// TIA Portal project "uppgift2" (V18)

(* hardware
DEVICE "S7-1500/ET200MP station_1"  S7-1500 station
   slot 0: "Rail_0"  Rack  6ES7 590-1***0-0AA0
   slot 1: "PLC_1"  CPU 1511C-1 PN  6ES7 511-1CK00-0AB0  V2.9
      slot 3: "CPU display_1"  6ES7591-1AA00-0AA0
      slot 32768: "PROFINET interface_1"  X1
         slot 32769: "Port_1"  X1 P1
         slot 32770: "Port_2"  X1 P2
      slot 34817: "Virtual CP interface port_1"  Virtual CP interface port  Virtual CP interface port
DEVICE "HMI_1"  KTP700 Mobile
   slot 0: "HMI_1"  KTP700 Mobile  6AV2 125-2GB03-0AX0  17.0.0.0
   slot 1: "HMI_RT_1"  KTP700 Mobile  6AV2 125-2GB03-0AX0  17.0.0.0
   slot 5: "HMI_1.IE_CP_1"  PROFINET Interface  17.0.0.0
      slot 1: "PROFINET Interface_1"  PROFINET Interface
         slot 1: "Port_1"  Port
*)

// ===== PLC "PLC_1"  CPU 1511C-1 PN =====

VAR_GLOBAL   // PLC tag table "Default tag table"
   "Start Button" AT %I0.0 : Bool;
   "Stop Button" AT %I0.1 : Bool;
   "Reset Button" AT %I0.2 : Bool;
   "Selective Mode" AT %I0.4 : Bool;
   "Base at place" AT %I0.5 : Bool;
   "Lid at place" AT %I0.6 : Bool;
   "Base is clamped" AT %I0.7 : Bool;
   "Lid is clamped" AT %I1.0 : Bool;
   "Item detected" AT %I1.1 : Bool;
   "Part is leaving (Sensor)" AT %I1.2 : Bool;
   "FACTORY I/O (Running)" AT %I1.3 : Bool;
   "Move X (Extend)" AT %Q0.0 : Bool;
   "Move Z (Lower)" AT %Q0.1 : Bool;
   "Grab Item" AT %Q0.2 : Bool;
   "Clamp base" AT %Q0.3 : Bool;
   "Clamp lid" AT %Q0.4 : Bool;
   "Lids emitter" AT %Q0.5 : Bool;
   "Lift Bases Clamp" AT %Q0.6 : Bool;
   "Lift Lids Clamp" AT %Q0.7 : Bool;
   "Counter" AT %QD30 : DInt;
   "Bases Vision Sensor" AT %ID30 : DInt;
   "Lids Vision Sensor" AT %ID34 : DInt;
   "Start Light" AT %Q1.0 : Bool;
   "Stop Light" AT %Q1.1 : Bool;
   "Reset Light" AT %Q1.2 : Bool;
   "Lids conveyor" AT %Q1.3 : Bool;
   "Bases conveyor" AT %Q1.4 : Bool;
   "Bases emitter" AT %Q1.5 : Bool;
   "flanker" AT %I2.4 : Bool;
   "Moving X (Sensor)" AT %I1.4 : Bool;
   "Moving Z (Sensor)" AT %I1.5 : Bool;
   "hmistop" AT %I2.2 : Bool;
   "hmireset" AT %I2.3 : Bool;
   "countyfinalflank" AT %I2.5 : Bool;
   "lids lift clamp limit" AT %I1.6 : Bool;
   "baselift clamp limit" AT %I1.7 : Bool;
   "countyflank" AT %I2.6 : Bool;
END_VAR

// folder: System blocks/Program resources

DATA_BLOCK "IEC_Timer_0_DB"   // DB3
{ S7_Optimized_Access := 'TRUE' }
AUTHOR : Simatic
FAMILY : IEC
NAME : IEC_TMR
VERSION : 1.0
// stored: InstanceOfName IEC_TIMER
"IEC_TIMER"
BEGIN
END_DATA_BLOCK

DATA_BLOCK "IEC_Timer_1_DB"   // DB4
{ S7_Optimized_Access := 'TRUE' }
AUTHOR : Simatic
FAMILY : IEC
NAME : IEC_TMR
VERSION : 1.0
// stored: InstanceOfName IEC_TIMER
"IEC_TIMER"
BEGIN
END_DATA_BLOCK

DATA_BLOCK "IEC_Counter_0_DB_2"   // DB5
{ S7_Optimized_Access := 'TRUE' }
AUTHOR : Simatic
FAMILY : IEC
NAME : CNTR
VERSION : 1.0
// stored: InstanceOfName IEC_COUNTER
"IEC_COUNTER"
BEGIN
END_DATA_BLOCK

DATA_BLOCK "IEC_Timer_0_DB_2"   // DB6
{ S7_Optimized_Access := 'TRUE' }
AUTHOR : Simatic
FAMILY : IEC
NAME : IEC_TMR
VERSION : 1.0
// stored: InstanceOfName IEC_TIMER
"IEC_TIMER"
BEGIN
END_DATA_BLOCK

DATA_BLOCK "IEC_Counter_0_DB_3"   // DB8
{ S7_Optimized_Access := 'TRUE' }
AUTHOR : Simatic
FAMILY : IEC
NAME : CNTR
VERSION : 1.0
// stored: InstanceOfName IEC_COUNTER
"IEC_COUNTER"
BEGIN
END_DATA_BLOCK

DATA_BLOCK "IEC_Counter_0_DB_4"   // DB10
{ S7_Optimized_Access := 'TRUE' }
AUTHOR : Simatic
FAMILY : IEC
NAME : CNTR
VERSION : 1.0
// stored: InstanceOfName IEC_COUNTER
"IEC_COUNTER"
BEGIN
END_DATA_BLOCK

DATA_BLOCK "IEC_Counter_0_DB_6"   // DB11
{ S7_Optimized_Access := 'TRUE' }
AUTHOR : Simatic
FAMILY : IEC
NAME : CNTR
VERSION : 1.0
// stored: InstanceOfName IEC_COUNTER
"IEC_COUNTER"
BEGIN
END_DATA_BLOCK

DATA_BLOCK "IEC_Counter_1_DB_1"   // DB12
{ S7_Optimized_Access := 'TRUE' }
AUTHOR : Simatic
FAMILY : IEC
NAME : CNTR
VERSION : 1.0
// stored: InstanceOfName IEC_COUNTER
"IEC_COUNTER"
BEGIN
END_DATA_BLOCK

DATA_BLOCK "IEC_Counter_0_DB_7"   // DB13
{ S7_Optimized_Access := 'TRUE' }
AUTHOR : Simatic
FAMILY : IEC
NAME : CNTR
VERSION : 1.0
// stored: InstanceOfName IEC_COUNTER
"IEC_COUNTER"
BEGIN
END_DATA_BLOCK

DATA_BLOCK "IEC_Counter_0_DB_5"   // DB14
{ S7_Optimized_Access := 'TRUE' }
AUTHOR : Simatic
FAMILY : IEC
NAME : CNTR
VERSION : 1.0
// stored: InstanceOfName IEC_COUNTER
"IEC_COUNTER"
BEGIN
END_DATA_BLOCK

DATA_BLOCK "IEC_Counter_0_DB_8"   // DB15
{ S7_Optimized_Access := 'TRUE' }
AUTHOR : Simatic
FAMILY : IEC
NAME : CNTR
VERSION : 1.0
// stored: InstanceOfName IEC_COUNTER
"IEC_COUNTER"
BEGIN
END_DATA_BLOCK

DATA_BLOCK "IEC_Counter_0_DB_9"   // DB16
{ S7_Optimized_Access := 'TRUE' }
AUTHOR : Simatic
FAMILY : IEC
NAME : CNTR
VERSION : 1.0
// stored: InstanceOfName IEC_COUNTER
"IEC_COUNTER"
BEGIN
END_DATA_BLOCK

DATA_BLOCK "IEC_Timer_5_DB"   // DB17
{ S7_Optimized_Access := 'TRUE' }
AUTHOR : Simatic
FAMILY : IEC
NAME : IEC_TMR
VERSION : 1.0
// stored: InstanceOfName IEC_TIMER
"IEC_TIMER"
BEGIN
END_DATA_BLOCK

DATA_BLOCK "IEC_Counter_0_DB"   // DB18
{ S7_Optimized_Access := 'TRUE' }
AUTHOR : Simatic
FAMILY : IEC
NAME : CNTR
VERSION : 1.0
// stored: InstanceOfName IEC_COUNTER
"IEC_COUNTER"
BEGIN
END_DATA_BLOCK

DATA_BLOCK "IEC_Timer_0_DB_4"   // DB20
{ S7_Optimized_Access := 'TRUE' }
AUTHOR : Simatic
FAMILY : IEC
NAME : IEC_TMR
VERSION : 1.0
// stored: InstanceOfName IEC_TIMER
"IEC_TIMER"
BEGIN
END_DATA_BLOCK

// folder: databases

DATA_BLOCK "outputs"   // DB1
{ S7_Optimized_Access := 'TRUE' }
VERSION : 0.1
   VAR
      RESETBUTTONHMI : Bool;
      Acutators : Struct
         "Move X (Extend)" : Bool;
         "Move Z (Lower)" : Bool;
         "Grab Item" : Bool;
         "Clamp base" : Bool;
         "Clamp lid" : Bool;
         "Lift Bases Clamp" : Bool;
         "Lift Lids Clamp" : Bool;
      END_STRUCT;
      BoxesCounters : Struct
         "green lids" : Int;
         "green bases" : Int;
         "blue lids" : Int;
         "blue bases" : Int;
         "bluegreen box" : Int;   // blå lock grön bas
         "greenblue box" : Int;   // grön bas blå lock
         "blue boxs" : Int;
         "green boxs" : Int;
         totalpartscounter : Int;
      END_STRUCT;
      Checks : Struct
         isreset : Bool;
         selectivestmode : Bool;
         pauseforselective : Bool;
      END_STRUCT;
      Modes : Struct
         "Run mode" : Bool;
         "Reset mode" : Bool;
         "Stop mode" : Bool;
      END_STRUCT;
      "Hmi-Producer" : Struct
         producedboxes : Int;
         toproduce : Int := 0;
      END_STRUCT;
   END_VAR
BEGIN
END_DATA_BLOCK

DATA_BLOCK "inputs"   // DB2
{ S7_Optimized_Access := 'TRUE' }
VERSION : 0.1
   VAR
      buttons : Struct
         "Start Button" : Bool;
         "Stop Button" : Bool;
         "Reset Button" : Bool;
      END_STRUCT;
      Sensors : Struct
         "Item detected" : Bool;
         "lid sensor value" : DInt;
      END_STRUCT;
      Sequences : Struct
         insequence : DInt;
         basesecquence : DInt;
         robotarmsequence : DInt;
      END_STRUCT;
      "green light" : Bool;
   END_VAR
BEGIN
END_DATA_BLOCK

DATA_BLOCK "functiondatabase"   // DB9
{ S7_Optimized_Access := 'TRUE' }
VERSION : 0.1
// stored: InstanceOfName hmi-order-limit&Color-total
"hmi-order-limit&Color-total"
BEGIN
END_DATA_BLOCK

DATA_BLOCK "tondb"   // DB19
{ S7_Optimized_Access := 'TRUE' }
VERSION : 0.1
   VAR
      IN : Bool;
      PT : Time := T#7000ms;
      Q : Bool;
      ET : Time;
   END_VAR
BEGIN
END_DATA_BLOCK

DATA_BLOCK "HMI-DB"   // DB1000
{ S7_Optimized_Access := 'TRUE' }
VERSION : 0.1
   VAR
      Inputs : Struct
         StartLight : Bool;
         StopLight : Bool;
         ResetLight : Bool;
      END_STRUCT;
      "Jogging&Priority" : Struct
         jogmode : Bool;
         hasbeenjogging : Bool;
         "jog bools" : Struct   // hmi jog bools
            "move x" : Bool;
            "move y" : Bool;
            "grab item" : Bool;
            "clamp lid" : Bool;
            "clamp base" : Bool;
            "lift base" : Bool;
            "lift lid" : Bool;
            "lid conv" : Bool;
            "base conv" : Bool;
            lampor : Bool;
         END_STRUCT;
         hmipriority : Bool;
         hmiprioritystate : Bool;
         resetdelivered : Bool;
      END_STRUCT;
   END_VAR
BEGIN
END_DATA_BLOCK

// folder: (top level)

FUNCTION_BLOCK "hmi-order-limit&Color-total"   // FB1, LAD
{ S7_Optimized_Access := 'TRUE' }
VERSION : 0.1
   VAR_OUTPUT
      basesadder : Int;
      lidadder : Int;
   END_VAR
BEGIN

REGION Network 1
   // limits the hmi to produce max 1000
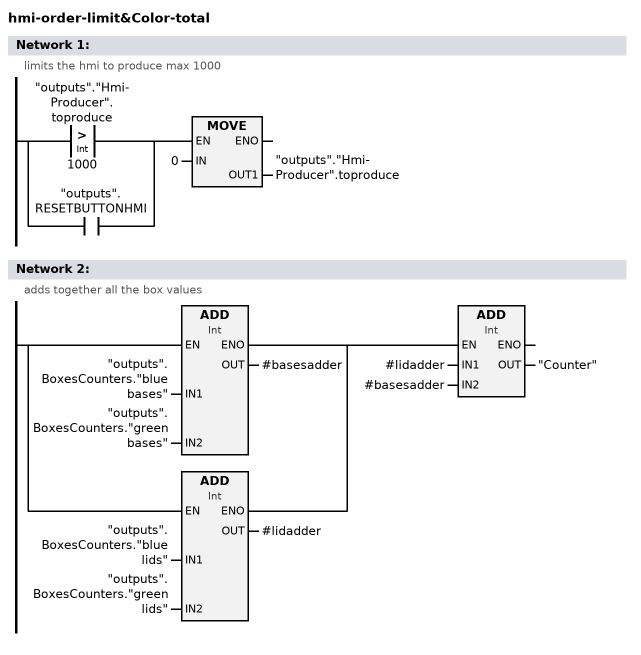
   RUNG wire#powerrail
      { S7_Templates := "SrcType := Int" } GT_Contact(in1 := "outputs"."Hmi-Producer".toproduce, in2 := 1000)
      wire#w1
      Move(in := 0, out1 => "outputs"."Hmi-Producer".toproduce)
   END_RUNG
   RUNG wire#powerrail
      Contact( "outputs".RESETBUTTONHMI )
   END_RUNG wire#w1
   // the same network as SCL:
   IF ("outputs"."Hmi-Producer".toproduce > 1000) OR "outputs".RESETBUTTONHMI THEN
       "outputs"."Hmi-Producer".toproduce := 0;
   END_IF;
END_REGION

REGION Network 2
   // adds together all the box values
   RUNG wire#powerrail
      { S7_Templates := "SrcType := Int" } Add(in1 := "outputs".BoxesCounters."blue bases", in2 := "outputs".BoxesCounters."green bases", out => #basesadder)
      wire#w1
      { S7_Templates := "SrcType := Int" } Add(in1 := #lidadder, in2 := #basesadder, out => "Counter")
   END_RUNG
   RUNG wire#powerrail
      { S7_Templates := "SrcType := Int" } Add(in1 := "outputs".BoxesCounters."blue lids", in2 := "outputs".BoxesCounters."green lids", out => #lidadder)
   END_RUNG wire#w1
   // the same network as SCL:
   #basesadder := "outputs".BoxesCounters."blue bases" + "outputs".BoxesCounters."green bases";
   #lidadder := "outputs".BoxesCounters."blue lids" + "outputs".BoxesCounters."green lids";
   IF TRUE OR TRUE THEN "Counter" := #lidadder + #basesadder; END_IF;
END_REGION
END_FUNCTION_BLOCK

FUNCTION "robotarm" : Void   // FC5, LAD
{ S7_Optimized_Access := 'TRUE' }
VERSION : 0.1
   VAR_TEMP   // added for the SCL form of the ladder/FBD networks
      _w1 : Bool;
   END_VAR
BEGIN

REGION Network 1
   // Both sequence 1 and 3 runs in the same network in an "or" statement, because both sequences need to use the "move z" acutator.
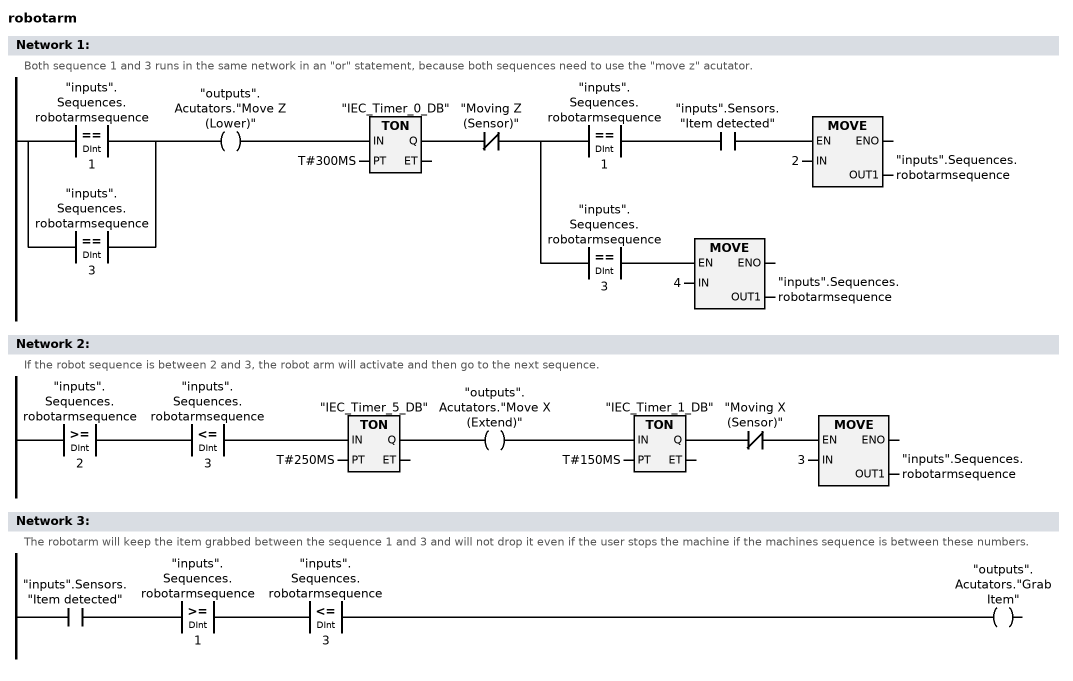
   "outputs".Acutators."Move Z (Lower)" := ("inputs".Sequences.robotarmsequence = 1) OR ("inputs".Sequences.robotarmsequence = 3);
   "IEC_Timer_0_DB".TON(IN := "outputs".Acutators."Move Z (Lower)", PT := T#300MS);
   #_w1 := "IEC_Timer_0_DB".Q AND NOT "Moving Z (Sensor)";
   IF #_w1 AND ("inputs".Sequences.robotarmsequence = 1) AND "inputs".Sensors."Item detected" THEN
       "inputs".Sequences.robotarmsequence := 2;
   END_IF;
   IF #_w1 AND ("inputs".Sequences.robotarmsequence = 3) THEN
       "inputs".Sequences.robotarmsequence := 4;
   END_IF;
END_REGION

REGION Network 2
   // If the robot sequence is between 2 and 3, the robot arm will activate and then go to the next sequence.
   "IEC_Timer_5_DB".TON(IN := ("inputs".Sequences.robotarmsequence >= 2) AND ("inputs".Sequences.robotarmsequence <= 3),
                        PT := T#250MS);
   "outputs".Acutators."Move X (Extend)" := "IEC_Timer_5_DB".Q;
   "IEC_Timer_1_DB".TON(IN := "IEC_Timer_5_DB".Q, PT := T#150MS);
   IF "IEC_Timer_1_DB".Q AND NOT "Moving X (Sensor)" THEN "inputs".Sequences.robotarmsequence := 3; END_IF;
END_REGION

REGION Network 3
   // The robotarm will keep the item grabbed between the sequence 1 and 3 and will not drop it even if the user stops the machine if the machines sequence is between these numbers.
   RUNG wire#powerrail
      Contact( "inputs".Sensors."Item detected" )
      { S7_Templates := "SrcType := DInt" } GE_Contact(in1 := "inputs".Sequences.robotarmsequence, in2 := 1)
      { S7_Templates := "SrcType := DInt" } LE_Contact(in1 := "inputs".Sequences.robotarmsequence, in2 := 3)
      Coil( "outputs".Acutators."Grab Item" )
   END_RUNG
   // the same network as SCL:
   "outputs".Acutators."Grab Item" := "inputs".Sensors."Item detected" AND ("inputs".Sequences.robotarmsequence >= 1) AND ("inputs".Sequences.robotarmsequence <= 3);
END_REGION
END_FUNCTION

FUNCTION "countcolors" : Void   // FC8, LAD
{ S7_Optimized_Access := 'TRUE' }
VERSION : 0.1
// This function counts the colors that passes through the colors sensors, both lid and base and then counts up accordingdly to which color that passed through the sensor.
   VAR_TEMP   // added for the SCL form of the ladder/FBD networks
      _w1 : Bool;
   END_VAR
BEGIN

REGION Network 1: counts final product
   // Counts the total boxes produced.
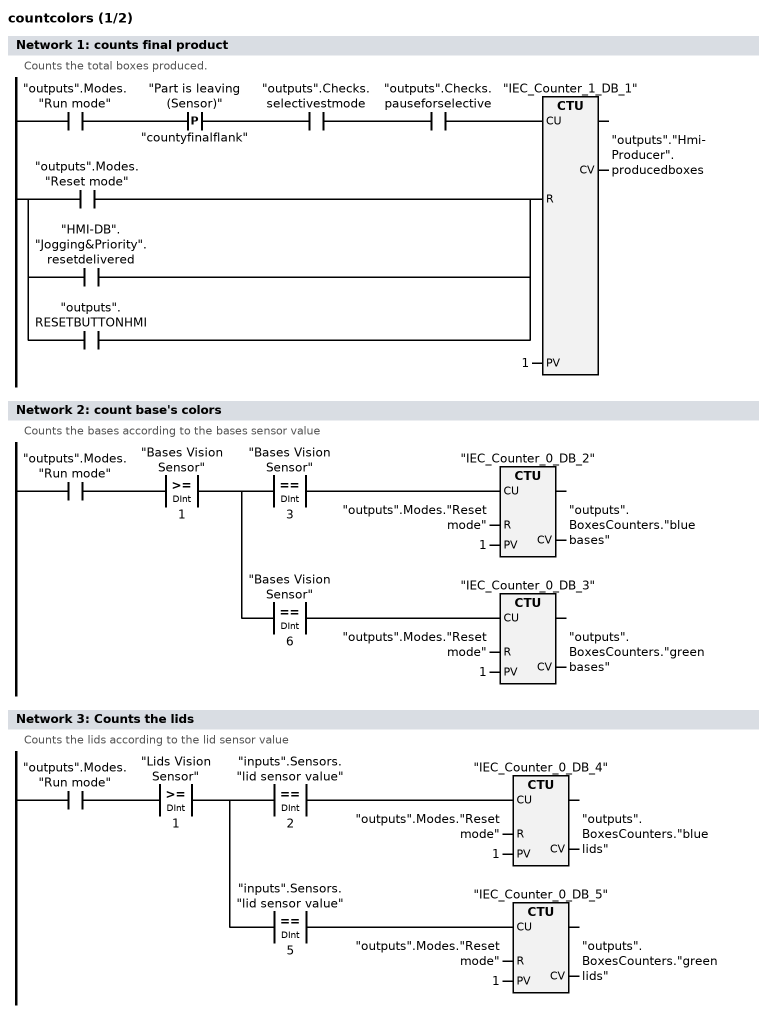
   #_w1 := "outputs".Modes."Run mode" AND "Part is leaving (Sensor)" AND NOT "countyfinalflank";   // rising edge of "Part is leaving (Sensor)"
   "countyfinalflank" := "Part is leaving (Sensor)";
   "IEC_Counter_1_DB_1".CTU(CU := #_w1 AND "outputs".Checks.selectivestmode AND "outputs".Checks.pauseforselective,
                           R := "outputs".Modes."Reset mode" OR "HMI-DB"."Jogging&Priority".resetdelivered OR "outputs".RESETBUTTONHMI,
                           PV := 1,
                           CV => "outputs"."Hmi-Producer".producedboxes);
END_REGION

REGION Network 2: count base's colors
   // Counts the bases according to the bases sensor value
   #_w1 := "outputs".Modes."Run mode" AND ("Bases Vision Sensor" >= 1);
   "IEC_Counter_0_DB_2".CTU(CU := #_w1 AND ("Bases Vision Sensor" = 3),
                           R := "outputs".Modes."Reset mode",
                           PV := 1,
                           CV => "outputs".BoxesCounters."blue bases");
   "IEC_Counter_0_DB_3".CTU(CU := #_w1 AND ("Bases Vision Sensor" = 6),
                           R := "outputs".Modes."Reset mode",
                           PV := 1,
                           CV => "outputs".BoxesCounters."green bases");
END_REGION

REGION Network 3: Counts the lids
   // Counts the lids according to the lid sensor value
   #_w1 := "outputs".Modes."Run mode" AND ("Lids Vision Sensor" >= 1);
   "IEC_Counter_0_DB_4".CTU(CU := #_w1 AND ("inputs".Sensors."lid sensor value" = 2),
                           R := "outputs".Modes."Reset mode",
                           PV := 1,
                           CV => "outputs".BoxesCounters."blue lids");
   "IEC_Counter_0_DB_5".CTU(CU := #_w1 AND ("inputs".Sensors."lid sensor value" = 5),
                           R := "outputs".Modes."Reset mode",
                           PV := 1,
                           CV => "outputs".BoxesCounters."green lids");
END_REGION

REGION Network 4
   // counts if the base and the lid is different colors
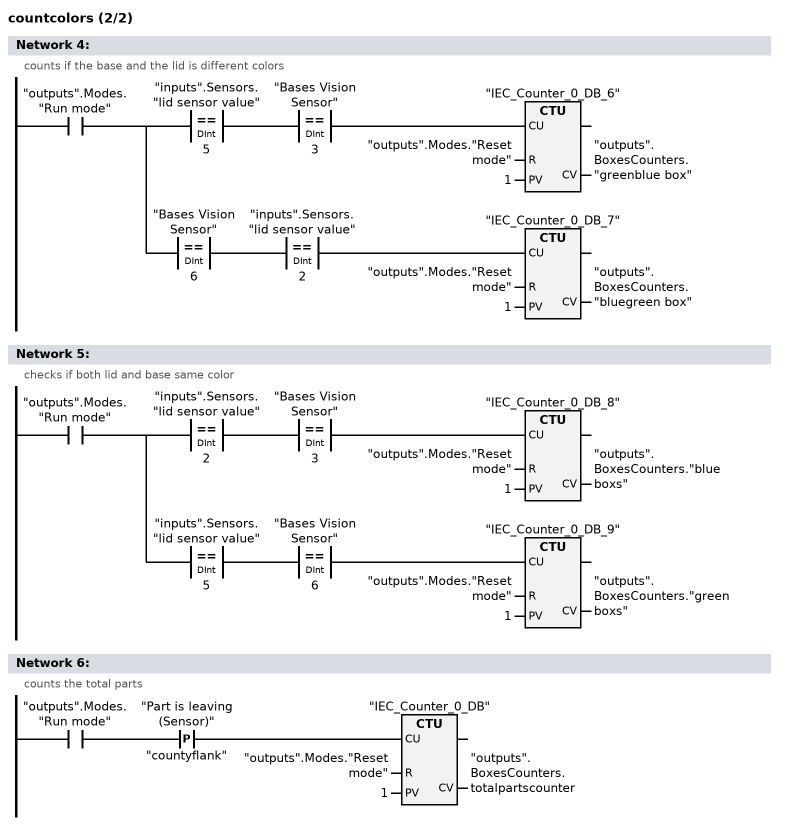
   "IEC_Counter_0_DB_6".CTU(CU := "outputs".Modes."Run mode" AND ("inputs".Sensors."lid sensor value" = 5) AND ("Bases Vision Sensor" = 3),
                           R := "outputs".Modes."Reset mode",
                           PV := 1,
                           CV => "outputs".BoxesCounters."greenblue box");
   "IEC_Counter_0_DB_7".CTU(CU := "outputs".Modes."Run mode" AND ("Bases Vision Sensor" = 6) AND ("inputs".Sensors."lid sensor value" = 2),
                           R := "outputs".Modes."Reset mode",
                           PV := 1,
                           CV => "outputs".BoxesCounters."bluegreen box");
END_REGION

REGION Network 5
   // checks if both lid and base same color
   "IEC_Counter_0_DB_8".CTU(CU := "outputs".Modes."Run mode" AND ("inputs".Sensors."lid sensor value" = 2) AND ("Bases Vision Sensor" = 3),
                           R := "outputs".Modes."Reset mode",
                           PV := 1,
                           CV => "outputs".BoxesCounters."blue boxs");
   "IEC_Counter_0_DB_9".CTU(CU := "outputs".Modes."Run mode" AND ("inputs".Sensors."lid sensor value" = 5) AND ("Bases Vision Sensor" = 6),
                           R := "outputs".Modes."Reset mode",
                           PV := 1,
                           CV => "outputs".BoxesCounters."green boxs");
END_REGION

REGION Network 6
   // counts the total parts
   #_w1 := "outputs".Modes."Run mode" AND "Part is leaving (Sensor)" AND NOT "countyflank";   // rising edge of "Part is leaving (Sensor)"
   "countyflank" := "Part is leaving (Sensor)";
   "IEC_Counter_0_DB".CTU(CU := #_w1,
                          R := "outputs".Modes."Reset mode",
                          PV := 1,
                          CV => "outputs".BoxesCounters.totalpartscounter);
END_REGION
END_FUNCTION

FUNCTION "resetscl" : Void   // FC9, SCL
{ S7_Optimized_Access := 'TRUE' }
VERSION : 0.1
BEGIN


   IF "outputs".Modes."Reset mode" THEN //Checks if its in reset mode
       "inputs".Sequences.basesecquence := 0; //Resets basesequence
       "inputs".Sequences.insequence := 0; //Resets lidsequence

       "tondb".IN := 1; 


       "IEC_Timer_0_DB_4".TON(IN := "tondb".IN, //Timer
                              PT := "tondb".PT,
                              Q => "tondb".Q,
                              ET => "tondb".ET);
       IF "tondb".Q THEN //When timer done then disable reset mode and set "isreset" variable to true
           "outputs".Checks.isreset := 1;
           "outputs".Modes."Reset mode" := 0;

           RESET_TIMER("IEC_Timer_0_DB_4");

       END_IF;

       IF NOT "Item detected" THEN //If arm not holding lid then reset the robot arm sequence
           "inputs".Sequences.robotarmsequence := 0;
       END_IF;

   END_IF;
END_FUNCTION

ORGANIZATION_BLOCK "Main"   // OB1, LAD, ProgramCycle
TITLE = "Main Program Sweep (Cycle)"
{ S7_Optimized_Access := 'TRUE' }
VERSION : 0.1
   VAR_INPUT
      Initial_Call : Bool;   // Initial call of this OB
      Remanence : Bool;   // =True, if remanent data are available
   END_VAR
BEGIN

REGION Network 1
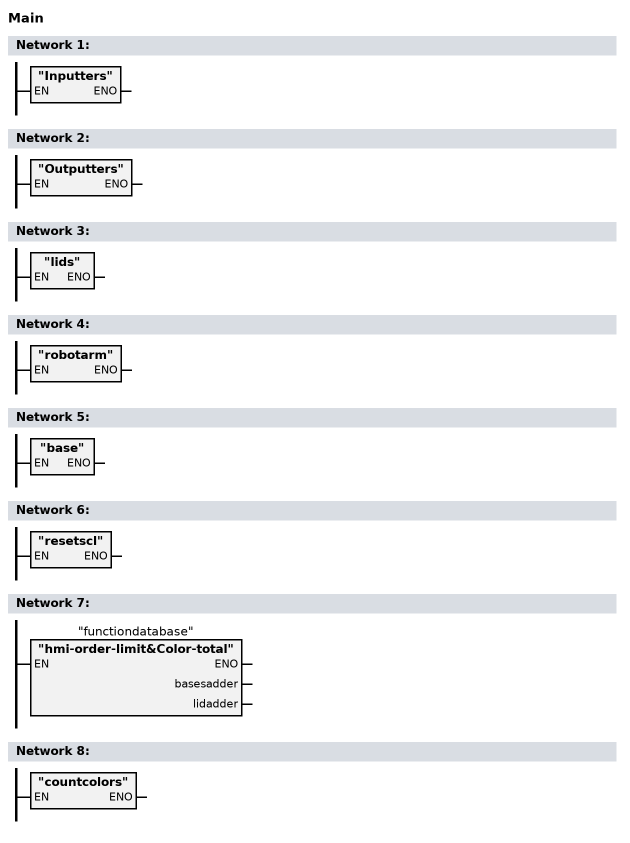
   RUNG wire#powerrail
      "Inputters"()
   END_RUNG
   // the same network as SCL:
   "Inputters"();
END_REGION

REGION Network 2
   RUNG wire#powerrail
      "Outputters"()
   END_RUNG
   // the same network as SCL:
   "Outputters"();
END_REGION

REGION Network 3
   RUNG wire#powerrail
      "lids"()
   END_RUNG
   // the same network as SCL:
   "lids"();
END_REGION

REGION Network 4
   RUNG wire#powerrail
      "robotarm"()
   END_RUNG
   // the same network as SCL:
   "robotarm"();
END_REGION

REGION Network 5
   RUNG wire#powerrail
      "base"()
   END_RUNG
   // the same network as SCL:
   "base"();
END_REGION

REGION Network 6
   RUNG wire#powerrail
      "resetscl"()
   END_RUNG
   // the same network as SCL:
   "resetscl"();
END_REGION

REGION Network 7
   RUNG wire#powerrail
      "functiondatabase"(basesadder =>, lidadder =>)
   END_RUNG
   // the same network as SCL:
   "functiondatabase"();   // "hmi-order-limit&Color-total"
END_REGION

REGION Network 8
   RUNG wire#powerrail
      "countcolors"()
   END_RUNG
   // the same network as SCL:
   "countcolors"();
END_REGION
END_ORGANIZATION_BLOCK

// folder: i/o

FUNCTION "Inputters" : Void   // FC1, LAD
{ S7_Optimized_Access := 'TRUE' }
VERSION : 0.1
   VAR_TEMP   // added for the SCL form of the ladder/FBD networks
      _w1 : Bool;
   END_VAR
BEGIN

REGION Network 1
   // if physical button is pressed then make the variables true
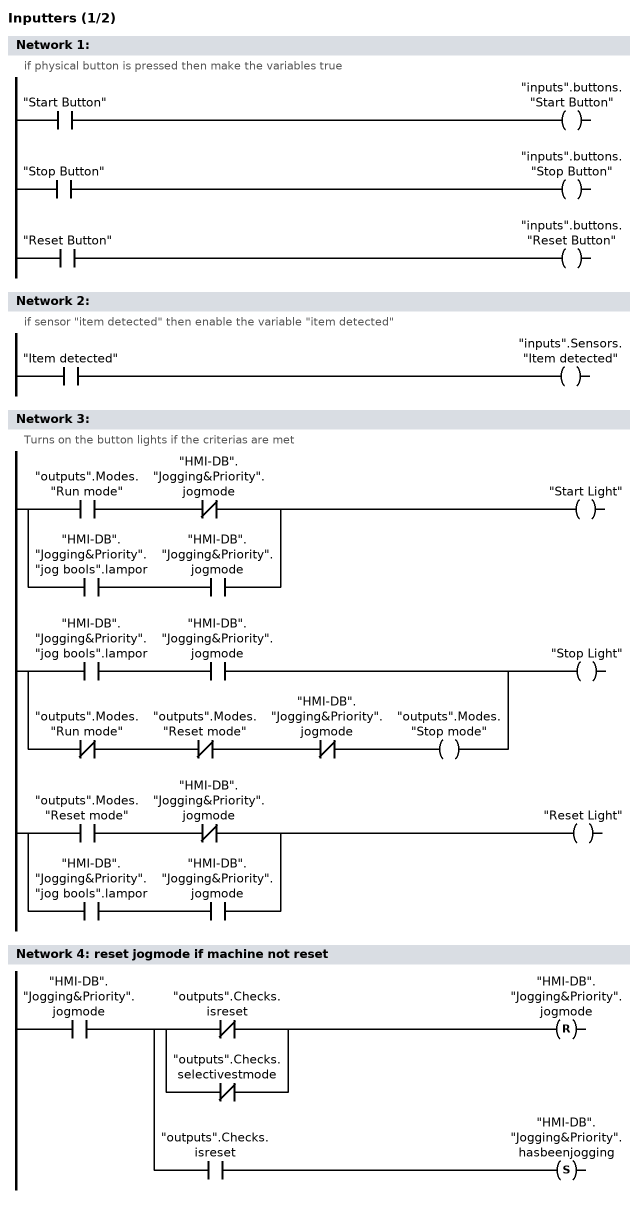
   RUNG wire#powerrail
      Contact( "Start Button" )
      Coil( "inputs".buttons."Start Button" )
   END_RUNG
   RUNG wire#powerrail
      Contact( "Stop Button" )
      Coil( "inputs".buttons."Stop Button" )
   END_RUNG
   RUNG wire#powerrail
      Contact( "Reset Button" )
      Coil( "inputs".buttons."Reset Button" )
   END_RUNG
   // the same network as SCL:
   "inputs".buttons."Start Button" := "Start Button";
   "inputs".buttons."Stop Button" := "Stop Button";
   "inputs".buttons."Reset Button" := "Reset Button";
END_REGION

REGION Network 2
   // if sensor "item detected" then enable the variable "item detected"
   RUNG wire#powerrail
      Contact( "Item detected" )
      Coil( "inputs".Sensors."Item detected" )
   END_RUNG
   // the same network as SCL:
   "inputs".Sensors."Item detected" := "Item detected";
END_REGION

REGION Network 3
   // Turns on the button lights if the criterias are met
   "Start Light" := ("outputs".Modes."Run mode" AND NOT "HMI-DB"."Jogging&Priority".jogmode) OR ("HMI-DB"."Jogging&Priority"."jog bools".lampor AND "HMI-DB"."Jogging&Priority".jogmode);
   "outputs".Modes."Stop mode" := NOT "outputs".Modes."Run mode" AND NOT "outputs".Modes."Reset mode" AND NOT "HMI-DB"."Jogging&Priority".jogmode;
   "Stop Light" := "outputs".Modes."Stop mode" OR ("HMI-DB"."Jogging&Priority"."jog bools".lampor AND "HMI-DB"."Jogging&Priority".jogmode);
   "Reset Light" := ("outputs".Modes."Reset mode" AND NOT "HMI-DB"."Jogging&Priority".jogmode) OR ("HMI-DB"."Jogging&Priority"."jog bools".lampor AND "HMI-DB"."Jogging&Priority".jogmode);
END_REGION

REGION Network 4: reset jogmode if machine not reset
   RUNG wire#powerrail
      Contact( "HMI-DB"."Jogging&Priority".jogmode )
      wire#w1
      I_Contact( "outputs".Checks.isreset )
      wire#w2
      R_Coil( "HMI-DB"."Jogging&Priority".jogmode )
   END_RUNG
   RUNG wire#w1
      I_Contact( "outputs".Checks.selectivestmode )
   END_RUNG wire#w2
   RUNG wire#w1
      Contact( "outputs".Checks.isreset )
      S_Coil( "HMI-DB"."Jogging&Priority".hasbeenjogging )
   END_RUNG
   // the same network as SCL:
   #_w1 := "HMI-DB"."Jogging&Priority".jogmode;
   IF "HMI-DB"."Jogging&Priority".jogmode AND (NOT "outputs".Checks.isreset OR NOT "outputs".Checks.selectivestmode) THEN
       "HMI-DB"."Jogging&Priority".jogmode := FALSE;
   END_IF;
   IF #_w1 AND "outputs".Checks.isreset THEN "HMI-DB"."Jogging&Priority".hasbeenjogging := TRUE; END_IF;
END_REGION

REGION Network 5
   // checks if the hmi is in priority mode and the hmi is in selective mode or that selective mode on the box is on
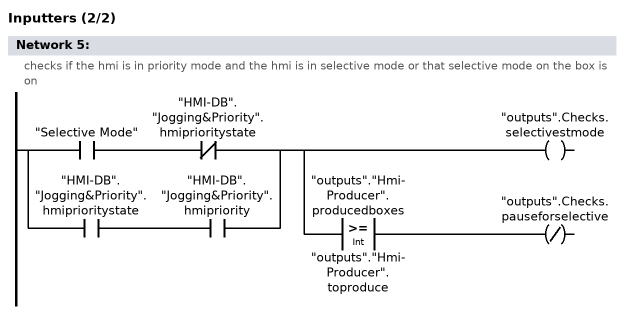
   RUNG wire#powerrail
      Contact( "Selective Mode" )
      I_Contact( "HMI-DB"."Jogging&Priority".hmiprioritystate )
      wire#w1
      Coil( "outputs".Checks.selectivestmode )
   END_RUNG
   RUNG wire#powerrail
      Contact( "HMI-DB"."Jogging&Priority".hmiprioritystate )
      Contact( "HMI-DB"."Jogging&Priority".hmipriority )
   END_RUNG wire#w1
   RUNG wire#w1
      { S7_Templates := "SrcType := Int" } GE_Contact(in1 := "outputs"."Hmi-Producer".producedboxes, in2 := "outputs"."Hmi-Producer".toproduce)
      I_Coil( "outputs".Checks.pauseforselective )
   END_RUNG
   // the same network as SCL:
   "outputs".Checks.selectivestmode := ("Selective Mode" AND NOT "HMI-DB"."Jogging&Priority".hmiprioritystate) OR ("HMI-DB"."Jogging&Priority".hmiprioritystate AND "HMI-DB"."Jogging&Priority".hmipriority);
   "outputs".Checks.pauseforselective := NOT ("outputs".Checks.selectivestmode AND ("outputs"."Hmi-Producer".producedboxes >= "outputs"."Hmi-Producer".toproduce));
END_REGION
END_FUNCTION

FUNCTION "Outputters" : Void   // FC2, LAD
{ S7_Optimized_Access := 'TRUE' }
VERSION : 0.1
   VAR_TEMP   // added for the SCL form of the ladder/FBD networks
      _w1 : Bool;
   END_VAR
BEGIN

REGION Network 1
   // Decides what mode should be enabled